      ProcessValue <- "F_Descargador_No"
   GraphicIOField "Campo ES gráfico_18" at 1195,401 size 28x28; PictureList "CheckBox"
      ProcessValue <- "F_Referencia_Menor_Descargador"
   IOField "Campo ES_7" at 1018,73 size 80x32; FormatPattern 9999999; Unit  mm
      ProcessValue <- "PosiciónEspera_F(Ant)"
   IOField "Campo ES_8" at 1018,97 size 80x32; FormatPattern 9999999; Unit  mm
      ProcessValue <- "PosiciónE1H1_F(Ant)"
   IOField "Campo ES_9" at 1018,121 size 80x32; FormatPattern 9999999; Unit  mm
      ProcessValue <- "PosiciónE1H2_F(Ant)"
   IOField "Campo ES_10" at 1018,145 size 80x32; FormatPattern 9999999; Unit  mm
      ProcessValue <- "PosiciónE2H1_F(Ant)"
   IOField "Campo ES_12" at 1018,169 size 80x32; FormatPattern 9999999; Unit  mm
      ProcessValue <- "PosiciónE2H2_F(Ant)"
   IOField "Campo ES_13" at 1018,193 size 80x32; FormatPattern 9999999; Unit  mm
      ProcessValue <- "PosiciónEntrega_F(Ant)"
   TextField "Campo de texto_34" at 249,678 size 130x18; Text 'DATOS PIEZA ACTUAL'
   TextField "Campo de texto_35" at 403,678 size 12x18; Text 'A'
   IOField "Champ E/S_24" at 414,675 size 53x25; FormatPattern 9999999
      ProcessValue <- "Pinza\Pinza.A"
      Appearance <- "Pinza\Pinza.PresenciaPieza"
   IOField "Champ E/S_25" at 483,675 size 53x25; FormatPattern 9999999
      ProcessValue <- "Pinza\Pinza.B"
      Appearance <- "Pinza\Pinza.PresenciaPieza"
   IOField "Champ E/S_26" at 554,675 size 53x24; FormatPattern 9999999
      ProcessValue <- "Pinza\Pinza.C"
      Appearance <- "Pinza\Pinza.PresenciaPieza"
   IOField "Champ E/S_27" at 629,675 size 53x25; FormatPattern 9999999
      ProcessValue <- "Pinza\Pinza.D"
      Appearance <- "Pinza\Pinza.PresenciaPieza"
   TextField "Campo de texto_36" at 472,678 size 11x18; Text 'B'
   TextField "Campo de texto_37" at 541,678 size 11x18; Text 'C'
   TextField "Campo de texto_38" at 616,678 size 12x18; Text 'D'
   TextField "Campo de texto_32" at 696,37 size 42x23; Text 'Pinza'
   TextField "Template_Plantilla_Campo de texto_4" at 696,67 size 568x3; Text 'Text'
   TextField "Template_Plantilla_Campo de texto_1" at 696,439 size 568x3; Text 'Text'
   TextField "Campo de texto_7" at 947,396 size 82x36; Text 'MOVIMIENTO SEGURO'
      Visibility <- "F_MovimientoSeguro"
      Appearance <- "F_MovimientoSeguro"
   TextField "Campo de texto_33" at 726,368 size 87x33; Text 'Tenaza Pleg. Atrás'
   TextField "Campo de texto_39" at 815,368 size 63x33; Text 'Herr. 1 OFF'
   TextField "Template_Plantilla_Campo de texto_3" at 696,359 size 568x3; Text 'Text'
   TextField "Campo de texto_43" at 882,368 size 63x33; Text 'Herr. 2 OFF'
   TextField "Campo de texto_18" at 1072,368 size 95x33; Text 'Descargador Atrás'
   TextField "Campo de texto_19" at 1160,368 size 95x33; Text 'Movimiento Corto'
   TextField "Campo de texto_10" at 719,242 size 191x25; Text 'Escalador relación mecánica'
   TextField "Campo de texto_13" at 719,262 size 191x25; Text 'Offset mecánico'
   TextField "Campo de texto_20" at 949,556 size 41x18; Text 'Martillo'
      Visibility <- "MANU"
   TextField "Campo de texto_23" at 825,556 size 35x18; Text 'Matriz'
      Visibility <- "MANU"
   TextField "Campo de texto_42" at 737,581 size 42x18; Text 'Herr. 1'
      Visibility <- "MANU"
   TextField "Campo de texto_45" at 737,622 size 42x18; Text 'Herr. 2'
      Visibility <- "MANU"
   TextField "Campo de texto_44" at 739,471 size 31x18; Text 'Pinza'
      Visibility <- "MANU"
   GraphicView "Visor de gráficos_1" at 1047,570 size 74x43; Picture "EMR2"
      Visibility <- "MANU"
   GraphicView "Visor de gráficos_2" at 1048,612 size 74x43; Picture "F1-3 EMR2"
      Visibility <- "MANU"
   GraphicView "Visor de gráficos_3" at 1152,612 size 74x43; Picture "F2-4 EMR2"
      Visibility <- "MANU"
   GraphicView "Visor de gráficos_4" at 1150,570 size 74x43; Picture "F1-3 EMR2"
      Visibility <- "MANU"
   GraphicView "Visor de gráficos_5" at 1126,590 size 12x12; Picture "outline_arrow_forward_ios_white_18dp"
      Visibility <- "MANU"
   GraphicView "Visor de gráficos_6" at 1135,590 size 12x12; Picture "outline_arrow_forward_ios_white_18dp"
      Visibility <- "MANU"
   GraphicView "Visor de gráficos_7" at 1126,632 size 12x12; Picture "outline_arrow_forward_ios_white_18dp"
      Visibility <- "MANU"
   GraphicView "Visor de gráficos_8" at 1135,632 size 12x12; Picture "outline_arrow_forward_ios_white_18dp"
      Visibility <- "MANU"
   TextField "Campo de texto_40" at 740,522 size 134x18; Text 'Bloque de Herramientas'
      Visibility <- "MANU"
   Button "Botón_42" at 48,625 size 40x40; TextOff 'Vista Condiciones'; PictureOff "Gráfico_7"
      on Click: ActivateScreen("eProC - 10 - Estados F_HW", 0)
   Button "Botón_11" at 1224,27 size 40x37; TextOff 'Vista Condiciones'; PictureOff "Tool"; Authorization "Nivel 3"
      on Click: ActivateScreen("eProC - 11 Referencias F-PL", 0)
   Button "Template_Plantilla_Bouton_2" at 1085,715 size 193x53; TextOff 'ALARMAS / DEFAUT'
      on Press: ActivateScreen("eProC - Alarmas", 0)
      Visibility <- "DB_OP.P_DEFAUT"

screen "eProC - 10 - Estados F_HW" 1280x768, template "Template"
   GraphicIOField "Campo ES gráfico_6" at 554,292 size 718x282; PictureList "Grupo 3 - Pinza1"
      ProcessValue <- "Alarma_Pinza"
   Polygon "Polígono_2" at 281,432 size 517x163
      Visibility <- "Pinza\Pinza.PresenciaPieza"
   Circle "Cercle_16" at 798,434 size 10x10
      Appearance <- "29S4"
   TextField "Campo de texto_29" at 910,349 size 114x18; Text '29S4 - Pinza Abierta'
   TextField "Campo de texto_30" at 894,313 size 116x18; Text '29S5 - Pinza Cerrada'
   Circle "Cercle_17" at 798,418 size 10x10
      Appearance <- "29S5"
   GraphicIOField "Campo ES gráfico_8" at 192,179 size 289x268; PictureList "Formador"
      ProcessValue <- "Alarma_Formador"
   Circle "Cercle_6" at 331,217 size 10x10
      Appearance <- "28S5"
   Circle "Cercle_7" at 331,246 size 10x10
      Appearance <- "28S6"
   TextField "Campo de texto_3" at 54,201 size 180x18; Text '28S5 - Herramientas Bloqueadas'
   TextField "Campo de texto_5" at 36,229 size 200x18; Text '28S6 - Herramientas Desbloqueadas'
   Circle "Cercle_8" at 406,291 size 10x10
      Appearance <- "28S3"
   Circle "Cercle_9" at 418,306 size 10x10
      Appearance <- "28S4"
   Circle "Cercle_10" at 460,360 size 10x10
      Appearance <- "28S1"
   Circle "Cercle_1" at 437,332 size 10x10
      Appearance <- "28S2"
   Circle "Cercle_0" at 371,397 size 10x10
      Appearance <- "27S5"
   Circle "Cercle_2" at 348,367 size 10x10
      Appearance <- "27S6"
   Circle "Cercle_18" at 313,326 size 10x10
      Appearance <- "27S7"
   Circle "Cercle_19" at 326,344 size 10x10
      Appearance <- "27S8"
   TextField "Campo de texto_10" at 488,240 size 146x18; Text '28S3 - Herr. 2 Matriz OFF'
   TextField "Campo de texto_15" at 496,267 size 142x18; Text '28S4 - Herr. 2 Matriz ON'
   TextField "Campo de texto_16" at 522,323 size 152x18; Text '28S1 - Herr. 2 Martillo OFF'
   TextField "Campo de texto_17" at 506,295 size 148x18; Text '28S2 - Herr. 2 Martillo ON'
   TextField "Campo de texto_11" at 44,381 size 146x18; Text '27S7 - Herr. 1 Matriz OFF'
   TextField "Campo de texto_19" at 46,411 size 142x18; Text '27S8 - Herr. 1 Matriz ON'
   TextField "Campo de texto_20" at 73,488 size 152x18; Text '27S5 - Herr. 1 Martillo OFF'
   TextField "Campo de texto_21" at 58,452 size 148x18; Text '27S6 - Herr. 1 Martillo ON'
   Button "Botón_42" at 48,625 size 40x40; TextOff 'Vista Condiciones'; PictureOff "Gráfico_6"
      on Click: ActivateScreen("eProC - 10 - Estados F", 0)
   TextField "Campo de texto_1" at 804,90 size 41x18; Text 'Martillo'
      Visibility <- "MANU"
   TextField "Campo de texto_23" at 680,90 size 35x18; Text 'Matriz'
      Visibility <- "MANU"
   TextField "Campo de texto_42" at 592,115 size 42x18; Text 'Herr. 1'
      Visibility <- "MANU"
   TextField "Campo de texto_45" at 592,156 size 42x18; Text 'Herr. 2'
      Visibility <- "MANU"
   TextField "Campo de texto_44" at 732,638 size 31x18; Text 'Pinza'
      Visibility <- "MANU"
   GraphicView "Visor de gráficos_1" at 904,108 size 74x43; Picture "EMR2"
      Visibility <- "MANU"
   GraphicView "Visor de gráficos_2" at 905,150 size 74x43; Picture "F1-3 EMR2"
      Visibility <- "MANU"
   GraphicView "Visor de gráficos_3" at 1009,150 size 74x43; Picture "F2-4 EMR2"
      Visibility <- "MANU"
   GraphicView "Visor de gráficos_4" at 1007,108 size 74x43; Picture "F1-3 EMR2"
      Visibility <- "MANU"
   GraphicView "Visor de gráficos_5" at 983,128 size 12x12; Picture "outline_arrow_forward_ios_white_18dp"
      Visibility <- "MANU"
   GraphicView "Visor de gráficos_6" at 992,128 size 12x12; Picture "outline_arrow_forward_ios_white_18dp"
      Visibility <- "MANU"
   GraphicView "Visor de gráficos_7" at 983,170 size 12x12; Picture "outline_arrow_forward_ios_white_18dp"
      Visibility <- "MANU"
   GraphicView "Visor de gráficos_8" at 992,170 size 12x12; Picture "outline_arrow_forward_ios_white_18dp"
      Visibility <- "MANU"
   TextField "Campo de texto_40" at 270,118 size 134x18; Text 'Bloque de Herramientas'
      Visibility <- "MANU"
   Button "Template_Plantilla_Bouton_2" at 1085,715 size 193x53; TextOff 'ALARMAS / DEFAUT'
      on Press: ActivateScreen("eProC - Alarmas", 0)
      Visibility <- "DB_OP.P_DEFAUT"
   TextField "Campo de texto_12" at 460,410 size 81x18; Text 'Herramienta 2'
   TextField "Campo de texto_13" at 366,434 size 81x18; Text 'Herramienta 1'
   Button "Botón_6" at 772,630 size 58x33; TextOff 'Avance'
      on Press: SetTag("DB_OP.RC2", 31); SetBit("DB_OP.OP_SELMANU2")
      Visibility <- "MANU"
      Appearance <- "DB_OP.RC2"
   Button "Botón_7" at 827,630 size 58x33; TextOff 'Retroc.'
      on Press: SetTag("DB_OP.RC2", 32); SetBit("DB_OP.OP_SELMANU2")
      Visibility <- "MANU"
      Appearance <- "DB_OP.RC2"
   Button "Botón_8" at 903,630 size 58x33; TextOff 'Abrir'
      on Press: SetTag("DB_OP.RC2", 33); SetBit("DB_OP.OP_SELMANU2")
      Visibility <- "MANU"
      Appearance <- "DB_OP.RC2"
   Button "Botón_9" at 959,630 size 58x33; TextOff 'Cerrar'
      on Press: SetTag("DB_OP.RC2", 34); SetBit("DB_OP.OP_SELMANU2")
      Visibility <- "MANU"
      Appearance <- "DB_OP.RC2"
   Button "Botón_34" at 496,110 size 58x33; TextOff 'Bajar'
      on Press: SetTag("DB_OP.RC2", 40); SetBit("DB_OP.OP_SELMANU2")
      Visibility <- "MANU"
      Appearance <- "DB_OP.RC2"
   Button "Botón_35" at 439,110 size 58x33; TextOff 'Subir'
      on Press: SetTag("DB_OP.RC2", 41); SetBit("DB_OP.OP_SELMANU2")
      Visibility <- "MANU"
      Appearance <- "DB_OP.RC2"
   Button "Botón_20" at 765,110 size 58x33; TextOff 'ON'
      on Press: SetTag("DB_OP.RC2", 42); SetBit("DB_OP.OP_SELMANU2")
      Visibility <- "MANU"
      Appearance <- "DB_OP.RC2"
   Button "Botón_21" at 765,149 size 58x33; TextOff 'ON'
      on Press: SetTag("DB_OP.RC2", 46); SetBit("DB_OP.OP_SELMANU2")
      Visibility <- "MANU"
      Appearance <- "DB_OP.RC2"
   Button "Botón_22" at 821,110 size 58x33; TextOff 'OFF'
      on Press: SetTag("DB_OP.RC2", 43); SetBit("DB_OP.OP_SELMANU2")
      Visibility <- "MANU"
      Appearance <- "DB_OP.RC2"
   Button "Botón_23" at 821,149 size 58x33; TextOff 'OFF'
      on Press: SetTag("DB_OP.RC2", 47); SetBit("DB_OP.OP_SELMANU2")
      Visibility <- "MANU"
      Appearance <- "DB_OP.RC2"
   Button "Botón_28" at 641,110 size 58x33; TextOff 'ON'
      on Press: SetTag("DB_OP.RC2", 44); SetBit("DB_OP.OP_SELMANU2")
      Visibility <- "MANU"
      Appearance <- "DB_OP.RC2"
   Button "Botón_5" at 641,148 size 58x33; TextOff 'ON'
      on Press: SetTag("DB_OP.RC2", 48); SetBit("DB_OP.OP_SELMANU2")
      Visibility <- "MANU"
      Appearance <- "DB_OP.RC2"
   Button "Botón_10" at 697,110 size 58x33; TextOff 'OFF'
      on Press: SetTag("DB_OP.RC2", 45); SetBit("DB_OP.OP_SELMANU2")
      Visibility <- "MANU"
      Appearance <- "DB_OP.RC2"
   Button "Botón_31" at 697,148 size 58x33; TextOff 'OFF'
      on Press: SetTag("DB_OP.RC2", 49); SetBit("DB_OP.OP_SELMANU2")
      Visibility <- "MANU"
      Appearance <- "DB_OP.RC2"

screen "eProC - 11 Referencias F-PL" 1280x768, template "Template"
   GraphicView "Visor de gráficos_1" at 134,72 size 979x505; Picture "Referencias"
   IOField "Champ E/S" at 340,310 size 80x27; Authorization "Nivel 2"; FormatPattern 9999999
      ProcessValue <- "Distancia_entre_Herramienta1_y_Pos0_F"
   IOField "Champ E/S_0" at 540,342 size 80x26; Authorization "Nivel 2"; FormatPattern 9999999
      ProcessValue <- "Distancia_entre_Pos0_y_Tenaza_F"
   TextField "Campo de texto_1" at 334,240 size 90x68; Text 'Distancia de Herramienta 1 a posición 0mm Pinza'
   TextField "Campo de texto_3" at 526,300 size 126x36; Text 'Distancia 0mm Pinza a Tenaza Plegadora'
   IOField "Champ E/S_2" at 552,526 size 80x26; Authorization "Nivel 2"; FormatPattern 9999999
      ProcessValue <- "Distancia_entre_Pos0_y_Descargador_F"
   TextField "Campo de texto_6" at 505,553 size 176x36; Text 'Distancia posición 0mm Pinza al Descargador'
   IOField "Champ E/S_3" at 235,566 size 80x27; Authorization "Nivel 2"; FormatPattern 9999999
      ProcessValue <- "Distancia_entre_Herramientas_F"
   TextField "Campo de texto_7" at 230,594 size 93x36; Text 'Distancia entre Herramientas'
   IOField "Champ E/S_4" at 592,610 size 80x26; Authorization "Nivel 2"; FormatPattern s9999999999
      ProcessValue <- "PosiciónMáxima_F"
   TextField "Campo de texto_8" at 587,636 size 93x36; Text 'Distancia Avance Máximo'
   IOField "Champ E/S_1" at 907,300 size 80x26; Authorization "Nivel 2"; FormatPattern 9999999
      ProcessValue <- "Distancia_entre_Pleg_Alin_PL"
   TextField "Campo de texto_2" at 861,330 size 196x20; Text 'Distancia de Plegador a Alineador'
   Switch "Interruptor_1" at 209,115 size 125x80; TextOn 'SI'; CaptionText 'Habilitar reglas'; TextOff 'NO'
      ProcessValue <- "HabilitarReglasBaluff"
   Button "Botón_1" at 440,76 size 135x50; TextOff 'Referenciar PL1'
      on Release: ResetBit("SolRef_PL1")
      on Press: SetBit("SolRef_PL1")
      Appearance <- "Homing_PL1"
      ObjectEnable <- "HabRefPleg"
      Visibility <- "HabRefPleg"
   Button "Botón_2" at 941,76 size 135x50; TextOff 'Referenciar PL2'
      on Release: ResetBit("SolRef_PL2")
      on Press: SetBit("SolRef_PL2")
      Appearance <- "Homing_PL2"
      ObjectEnable <- "HabRefPleg"
      Visibility <- "HabRefPleg"
   Button "Template_Plantilla_Bouton_2" at 1085,715 size 193x53; TextOff 'ALARMAS / DEFAUT'
      on Press: ActivateScreen("eProC - Alarmas", 0)
      Visibility <- "DB_OP.P_DEFAUT"

screen "eProC - Recetas" 1280x768, template "Template"
   IOField "Champ E/S_43" at 357,162 size 98x23; FormatPattern 9999999; Unit  mm
      ProcessValue <- "Receta\Recetas.B"
   IOField "Champ E/S_44" at 869,304 size 90x23; FormatPattern 9999999; Unit  mm
      ProcessValue <- "Receta\Recetas.C"
   IOField "Champ E/S_46" at 743,113 size 96x24; FormatPattern s999999; Unit  mm
      ProcessValue <- "Receta\Recetas.F2"
   IOField "Champ E/S_47" at 743,90 size 90x23; FormatPattern s999999; Unit  mm
      ProcessValue <- "Receta\Recetas.F1"
   IOField "Champ E/S_48" at 561,90 size 94x23; FormatPattern s999999; Unit  mm
      ProcessValue <- "Receta\Recetas.F3"
   IOField "Champ E/S_49" at 581,137 size 96x24; FormatPattern s999999; Unit  mm
      ProcessValue <- "Receta\Recetas.PL1_2"
   IOField "Champ E/S_50" at 193,137 size 91x24; FormatPattern s999999; Unit  mm
      ProcessValue <- "Receta\Recetas.PL1_1"
   IOField "Champ E/S_51" at 1165,137 size 94x24; FormatPattern s999999; Unit  mm
      ProcessValue <- "Receta\Recetas.PL2_1"
   TextField "Campo de texto_56" at 340,160 size 17x26; Text 'B'
   TextField "Campo de texto_57" at 852,302 size 17x26; Text 'C'
   IOField "Champ E/S_52" at 1121,303 size 88x24; FormatPattern 9999999; Unit  mm
      ProcessValue <- "Receta\Recetas.D"
   TextField "Campo de texto_60" at 1103,302 size 19x26; Text 'D'
   IOField "Champ E/S_53" at 561,112 size 94x25; FormatPattern s999999; Unit  mm
      ProcessValue <- "Receta\Recetas.F4"
   IOField "Champ E/S_54" at 764,137 size 93x24; FormatPattern s999999; Unit  mm
      ProcessValue <- "Receta\Recetas.PL2_2"
   TextField "Campo de texto_62" at 556,302 size 17x26; Text 'A'
   IOField "Champ E/S_55" at 575,304 size 94x23; FormatPattern 9999999; Unit  mm
      ProcessValue <- "Receta\Recetas.A"
   TextField "Campo de texto_63" at 542,138 size 40x22; Text 'PL1-2'
   TextField "Campo de texto_64" at 726,113 size 20x22; Text 'F2'
   TextField "Campo de texto_65" at 152,138 size 40x22; Text 'PL1-1'
   TextField "Campo de texto_66" at 726,89 size 20x22; Text 'F1'
   TextField "Campo de texto_67" at 725,138 size 40x22; Text 'PL2-2'
   TextField "Campo de texto_68" at 541,113 size 20x22; Text 'F4'
   TextField "Campo de texto_69" at 1124,138 size 40x22; Text 'PL2-1'
   TextField "Campo de texto_70" at 541,89 size 20x22; Text 'F3'
   RecipeView "RecipeView" at 25,65 size 307x64; RecipeNameCaption 'Receta:'; DataRecordNameCaption 'Receta:'; ValueCaption 'Valor'; RecipeNrCaption 'N.º:'; DataRecordNrCaption 'Nº:'; EntryNameCaption 'Nombre de entrada'; Recipe "Pieza"; Tag4DataRecord "Receta\Recetas.Nombre"
   Button "Button_7" at 856,371 size 82x33; TextOff 'Cargar'; PictureOff "Flèche_Droite"
      on Press: SetBit("Receta\Recetas.x_M2"); function_eba64363('REFERENCE', "Receta\Recetas.Nombre", 1, N)
      Appearance <- "Receta\Recetas.x_M2"
   TextField "Campo de texto_15" at 953,376 size 72x22; Text 'Almacén 2'
   IOField "Champ E/S_57" at 1041,376 size 118x24; FormatPattern ????????????????????
      ProcessValue <- "Almacén 2\PAlmacén.Nombre"
   TextField "Campo de texto_59" at 39,37 size 159x26; Text 'Selección de Receta'
   Button "Button_6" at 42,368 size 82x35; TextOff 'Cargar'; PictureOff "Flèche_Droite"
      on Press: SetBit("Receta\Recetas.x_M1"); function_eba64363('REFERENCE', "Receta\Recetas.Nombre", 1, N)
      Appearance <- "Receta\Recetas.x_M1"
   TextField "Campo de texto_14" at 139,375 size 72x22; Text 'Almacén 1'
   IOField "Champ E/S_56" at 227,375 size 120x24; FormatPattern ????????????????????
      ProcessValue <- "Almacén 1\PAlmacén.Nombre"
   IOField "Champ E/S_1" at 289,304 size 90x23; FormatPattern 9999999; Unit  mm
      ProcessValue <- "Receta\Recetas.C"
   TextField "Campo de texto_1" at 272,302 size 17x26; Text 'C'
   IOField "Champ E/S_2" at 41,303 size 88x24; FormatPattern 9999999; Unit  mm
      ProcessValue <- "Receta\Recetas.D"
   TextField "Campo de texto_2" at 23,302 size 19x26; Text 'D'
   Button "Template_Plantilla_Bouton_1" at 345,50 size 150x63; TextOff 'EDITAR RECETAS / SYSTEM'; Authorization "Nivel 3"
      on Click: ActivateScreen("eProC - Edición Recetas", 0)
   Button "Template_Plantilla_Botón_32" at 129,715 size 150x53; TextOff 'SELECCIÓN RECETAS'
   Button "Template_Plantilla_Bouton_2" at 1085,715 size 193x53; TextOff 'ALARMAS / DEFAUT'
      on Press: ActivateScreen("eProC - Alarmas", 0)
      Visibility <- "DB_OP.P_DEFAUT"
   IOField "Campo ES_1" at 321,415 size 130x34; FormatPattern 9999999999
      ProcessValue <- "Descargador-ID_Bobina_Alm1"
   IOField "Campo ES_2" at 1136,415 size 130x34; FormatPattern 9999999999
      ProcessValue <- "Descargador-ID_Bobina_Alm2"
   DateTimeField "Campo de fecha y hora_1" at 180,415 size 131x34
      ProcessValue <- "Descargador-FechaCorte_Alm1"
   DateTimeField "Campo de fecha y hora_2" at 995,415 size 131x34
      ProcessValue <- "Descargador-FechaCorte_Alm2"
   SymbolicIOField "Campo ES simbólico_1" at 41,415 size 130x34; TextOff '0'; TextOn '1'; TextList "Proveedor"
      ProcessValue <- "Proveedor_Indexado_Alm1"
   SymbolicIOField "Campo ES simbólico_2" at 856,415 size 130x34; TextOff '0'; TextOn '1'; TextList "Proveedor"
      ProcessValue <- "Proveedor_Indexado_Alm2"
   IOField "Champ E/S_74" at 302,520 size 64x32; Authorization "Nivel 1"; FormatPattern s999999; Unit   
      ProcessValue <- "Almacén 1\PAlmacén.F2"
   IOField "Champ E/S_75" at 302,493 size 64x32; Authorization "Nivel 1"; FormatPattern s999999; Unit   
      ProcessValue <- "Almacén 1\PAlmacén.F1"
   IOField "Champ E/S_76" at 86,498 size 64x32; Authorization "Nivel 1"; FormatPattern s999999; Unit   
      ProcessValue <- "Almacén 1\PAlmacén.F3"
   IOField "Champ E/S_77" at 86,471 size 64x32; Authorization "Nivel 1"; FormatPattern s999999; Unit   
      ProcessValue <- "Almacén 1\PAlmacén.PL1_2"
   IOField "Champ E/S_78" at 86,648 size 64x32; Authorization "Nivel 1"; FormatPattern s999999; Unit   
      ProcessValue <- "Almacén 1\PAlmacén.PL1_1"
   IOField "Champ E/S_79" at 302,651 size 64x32; Authorization "Nivel 1"; FormatPattern s999999; Unit   
      ProcessValue <- "Almacén 1\PAlmacén.PL2_1"
   IOField "Champ E/S_81" at 86,525 size 64x32; Authorization "Nivel 1"; FormatPattern s999999; Unit   
      ProcessValue <- "Almacén 1\PAlmacén.F4"
   IOField "Champ E/S_82" at 302,466 size 64x32; Authorization "Nivel 1"; FormatPattern s999999; Unit   
      ProcessValue <- "Almacén 1\PAlmacén.PL2_2"
   TextField "Campo de texto_80" at 46,476 size 40x22; Text 'PL1-2'
   TextField "Campo de texto_81" at 366,526 size 20x22; Text 'F2'
   TextField "Campo de texto_82" at 46,652 size 40x22; Text 'PL1-1'
   TextField "Campo de texto_83" at 366,497 size 20x22; Text 'F1'
   TextField "Campo de texto_84" at 364,471 size 40x22; Text 'PL2-2'
   TextField "Campo de texto_85" at 66,531 size 20x22; Text 'F4'
   TextField "Campo de texto_86" at 364,655 size 40x22; Text 'PL2-1'
   TextField "Campo de texto_87" at 66,502 size 20x22; Text 'F3'
   IOField "Champ E/S_15" at 904,498 size 64x32; Authorization "Nivel 1"; FormatPattern s999999; Unit   
      ProcessValue <- "Almacén 2\PAlmacén.F3"
   IOField "Champ E/S_16" at 904,471 size 64x32; Authorization "Nivel 1"; FormatPattern s999999; Unit   
      ProcessValue <- "Almacén 2\PAlmacén.PL1_2"
   IOField "Champ E/S_58" at 904,648 size 65x32; Authorization "Nivel 1"; FormatPattern s999999; Unit   
      ProcessValue <- "Almacén 2\PAlmacén.PL1_1"
   IOField "Champ E/S_60" at 904,525 size 64x32; Authorization "Nivel 1"; FormatPattern s999999; Unit   
      ProcessValue <- "Almacén 2\PAlmacén.F4"
   TextField "Campo de texto_53" at 865,476 size 40x22; Text 'PL1-2'
   TextField "Campo de texto_55" at 865,652 size 40x22; Text 'PL1-1'
   TextField "Campo de texto_58" at 885,531 size 20x22; Text 'F4'
   TextField "Campo de texto_7" at 885,502 size 20x22; Text 'F3'
   IOField "Champ E/S_13" at 1119,520 size 64x32; Authorization "Nivel 1"; FormatPattern s999999; Unit   
      ProcessValue <- "Almacén 2\PAlmacén.F2"
   IOField "Champ E/S_14" at 1119,493 size 64x32; Authorization "Nivel 1"; FormatPattern s999999; Unit   
      ProcessValue <- "Almacén 2\PAlmacén.F1"
   IOField "Champ E/S_59" at 1119,651 size 64x32; Authorization "Nivel 1"; FormatPattern s999999; Unit   
      ProcessValue <- "Almacén 2\PAlmacén.PL2_1"
   IOField "Champ E/S_61" at 1119,466 size 64x32; Authorization "Nivel 1"; FormatPattern s999999; Unit   
      ProcessValue <- "Almacén 2\PAlmacén.PL2_2"
   TextField "Campo de texto_54" at 1180,526 size 20x22; Text 'F2'
   TextField "Campo de texto_4" at 1180,497 size 20x22; Text 'F1'
   TextField "Campo de texto_5" at 1180,471 size 40x22; Text 'PL2-2'
   TextField "Campo de texto_6" at 1180,655 size 40x22; Text 'PL2-1'
   IOField "Champ E/S_3" at 86,581 size 64x32; Authorization "Nivel 1"; FormatPattern s999999; Unit   
      ProcessValue <- "Almacén 1\PAlmacén.C"
   TextField "Campo de texto_3" at 66,587 size 13x22; Text 'C'
   IOField "Champ E/S_4" at 904,581 size 64x32; Authorization "Nivel 1"; FormatPattern s999999; Unit   
      ProcessValue <- "Almacén 2\PAlmacén.C"
   TextField "Campo de texto_8" at 885,587 size 13x22; Text 'C'

screen "eProC - Defectos" 1280x768, template "Template"
   TextField "Campo de texto_14" at 18,389 size 97x28; Text 'Almacén 2'
   TextField "Campo de texto_7" at 693,45 size 95x28; Text 'Esquina 1'
   TextField "Campo de texto_8" at 532,45 size 95x28; Text 'Esquina 2'
   TextField "Campo de texto_9" at 364,97 size 138x28; Text 'Herramienta 1'
   TextField "Campo de texto_10" at 364,154 size 138x28; Text 'Herramienta 2'
   TextField "Campo de texto_2" at 982,66 size 85x28; Text 'Contador'
   TextField "Campo de texto_1" at 18,45 size 97x28; Text 'Almacén 1'
   TextField "Campo de texto_3" at 693,381 size 90x28; Text 'Esquina 1'
   TextField "Campo de texto_4" at 532,381 size 90x28; Text 'Esquina 2'
   TextField "Campo de texto_5" at 364,433 size 133x28; Text 'Herramienta 1'
   TextField "Campo de texto_6" at 364,490 size 133x28; Text 'Herramienta 2'
   TextField "Campo de texto_16" at 982,402 size 85x28; Text 'Contador'
   TextField "Campo de texto_11" at 316,306 size 102x28; Text 'Plegadores'
   TextField "Campo de texto_12" at 316,642 size 102x28; Text 'Plegadores'
   Button "Template_Plantilla_Botón_55" at 789,715 size 150x53; TextOff 'ACUSAR DEFECTO'
   IOField "Campo ES_1" at 980,106 size 96x32; FormatPattern 9999
      ProcessValue <- "Contador_def_Alm1"
   Button "Botón_1" at 520,92 size 120x40; TextOff 'E2 H1'
      on Click: function_dd21b452("Contador_def_Alm1", 1); SetTag("Defecto_Alm1", 3)
   Button "Botón_2" at 680,92 size 120x40; TextOff 'E1 H1'
      on Click: function_dd21b452("Contador_def_Alm1", 1); SetTag("Defecto_Alm1", 1)
   Button "Botón_3" at 520,148 size 120x40; TextOff 'E2 H2'
      on Click: function_dd21b452("Contador_def_Alm1", 1); SetTag("Defecto_Alm1", 4)
   Button "Botón_4" at 680,148 size 120x40; TextOff 'E1 H2'
      on Click: function_dd21b452("Contador_def_Alm1", 1); SetTag("Defecto_Alm1", 2)
   Button "Botón_5" at 472,300 size 120x40; TextOff 'PL1-2'
      on Click: function_dd21b452("Contador_def_Alm1", 1); SetTag("Defecto_Alm1", 5)
   Button "Botón_6" at 632,300 size 120x40; TextOff 'PL2-2'
      on Click: function_dd21b452("Contador_def_Alm1", 1); SetTag("Defecto_Alm1", 6)
   Button "Botón_7" at 980,146 size 120x40; TextOff 'Reset'
      on Click: SetTag("Contador_def_Alm1", 0)
   IOField "Campo ES_2" at 980,442 size 96x32; FormatPattern 9999
      ProcessValue <- "Contador_def_Alm2"
   Button "Botón_8" at 520,428 size 120x40; TextOff 'E2 H1'
      on Click: function_dd21b452("Contador_def_Alm2", 1); SetTag("Defecto_Alm2", 3)
   Button "Botón_9" at 680,428 size 120x40; TextOff 'E1 H1'
      on Click: function_dd21b452("Contador_def_Alm2", 1); SetTag("Defecto_Alm2", 1)
   Button "Botón_10" at 520,484 size 120x40; TextOff 'E2 H2'
      on Click: function_dd21b452("Contador_def_Alm2", 1); SetTag("Defecto_Alm2", 4)
   Button "Botón_11" at 680,484 size 120x40; TextOff 'E1 H2'
      on Click: function_dd21b452("Contador_def_Alm2", 1); SetTag("Defecto_Alm2", 2)
   Button "Botón_12" at 472,636 size 120x40; TextOff 'PL1-2'
      on Click: function_dd21b452("Contador_def_Alm2", 1); SetTag("Defecto_Alm2", 5)
   Button "Botón_13" at 632,636 size 120x40; TextOff 'PL2-2'
      on Click: function_dd21b452("Contador_def_Alm2", 1); SetTag("Defecto_Alm2", 6)
   Button "Botón_14" at 980,482 size 120x40; TextOff 'Reset'
      on Click: SetTag("Contador_def_Alm2", 0)
   Button "Template_Plantilla_Bouton_2" at 1085,715 size 193x53; TextOff 'ALARMAS / DEFAUT'
      on Press: ActivateScreen("eProC - Alarmas", 0)
      Visibility <- "DB_OP.P_DEFAUT"
   IOField "Champ E/S_1" at 122,392 size 171x24; FormatPattern ????????????????????
      ProcessValue <- "Almacén 2\PAlmacén.Nombre"
   IOField "Champ E/S_2" at 122,48 size 170x24; FormatPattern ????????????????????
      ProcessValue <- "Almacén 1\PAlmacén.Nombre"

VB script "Script_1"
   'NOTE : Appuyez sur <Ctrl><Espacement> pour lancer le script et afficher le large éventail de fonctions.
   'Ecrivez vos scripts en utilisant les fonctions système ou le modèle d'objet. Vous pouvez facilement accéder au
   'système via l'objet runtime IHM. Pour sélectionner rapidement une référence objet
   'vous pouvez appuyer sur <Alt><Flèche droite>. Vous pouvez créer des scripts complexes en ayant recours au
   'langage de programmation VBScript et accéder directement aux variables via le nom, par ex. tag = 5.
*)

(* ===== HMI "HMI_RT_2" =====
system functions are stored by id; their names below are inferred from use
connection "HMI_ServidorHTTP": Web, WebPanel

HMI tags "Tabla de variables estándar"
   "Descargador-PiezaPresente" : Bool AT Descargador-PiezaPresente, 1 s   // Unidad presente en el descargador (DB12DBX46.0)
   "31S1 (E8.0)" : Bool AT 31S1, 1 s   // Presencia Producto en Descargador
      on ChangeValue: "FuncionVB_1"()
   "Evento_ArchivarVariable_1" : Bool, internal   // Para guardar los datos del producto en almacen 1
      on ChangeValue: function_abcfba0d("Cota C_Alm1"); function_abcfba0d("Factor F1_Alm1"); function_abcfba0d("Factor F2_Alm1"); function_abcfba0d("Factor F3_Alm1"); function_abcfba0d("Factor F4_Alm1"); function_abcfba0d("Factor PL1-1_Alm1"); function_abcfba0d("Factor PL1-2_Alm1"); function_abcfba0d("Factor PL2-1_Alm1"); function_abcfba0d("Factor PL2-2_Alm1"); function_abcfba0d("ID_Proveedor_Alm1"); function_abcfba0d("ID_FechaCorte_Alm1"); function_abcfba0d("ID_Bobina_Alm1")
   "Evento_ArchivarVariable_2" : Bool, internal   // Para guardar lel posicionamiento de la pinza en almacen 1
      on ChangeValue: function_abcfba0d("PosReal_E1H1_Alm1"); function_abcfba0d("PosReal_E1H2_Alm1"); function_abcfba0d("PosReal_E2H1_Alm1"); function_abcfba0d("PosReal_E2H2_Alm1"); function_abcfba0d("PosReal_Entrega_Alm1"); function_abcfba0d("PosReal_Recepcion_Alm1"); function_abcfba0d("Consigna_E1H1_Alm1"); function_abcfba0d("Consigna_E1H2_Alm1"); function_abcfba0d("Consigna_E2H1_Alm1"); function_abcfba0d("Consigna_E2H2_Alm1"); function_abcfba0d("Consigna_Entrega_Alm1"); function_abcfba0d("Consigna_Recepcion_Alm1")
   "Evento_ArchivarVariable_3" : Bool, internal   // Para guardar el posicionamiento de los plegadores en almacen 1
      on ChangeValue: function_abcfba0d("PosiciónEntrega_PL1_A1"); function_abcfba0d("PosiciónEspera_PL1_A1"); function_abcfba0d("PosiciónPlegado1_PL1_A1"); function_abcfba0d("PosiciónPlegado2_PL1_A1"); function_abcfba0d("PosiciónRecepción_PL1_A1"); function_abcfba0d("PosiciónEntrega_PL2_A1"); function_abcfba0d("PosiciónEspera_PL2_A1"); function_abcfba0d("PosiciónPlegado1_PL2_A1"); function_abcfba0d("PosiciónPlegado2_PL2_A1"); function_abcfba0d("PosiciónRecepción_PL2_A1")
   "Descargador-Almacen" : Bool AT Descargador-Almacen, 1 s   // Si este bit es 0 la unidad proviene del almacén 1, si vale 1 del almacén 2 (DB12DBX46.1)
   "Evento_ArchivarVariable_4" : Bool, internal   // Para guardar los datos del producto en almacen 2
      on ChangeValue: function_abcfba0d("Cota C_Alm2"); function_abcfba0d("Factor F1_Alm2"); function_abcfba0d("Factor F2_Alm2"); function_abcfba0d("Factor F3_Alm2"); function_abcfba0d("Factor F4_Alm2"); function_abcfba0d("Factor PL1-1_Alm2"); function_abcfba0d("Factor PL1-2_Alm2"); function_abcfba0d("Factor PL2-1_Alm2"); function_abcfba0d("Factor PL2-2_Alm2"); function_abcfba0d("ID_Prov_Ind_Alm2"); function_abcfba0d("ID_FechaCorte_Alm2"); function_abcfba0d("ID_Bobina_Alm2")
   "Aux1" : Bool, internal   // utilizada en FuncionVB_1
   "Aux2" : Bool, internal   // para entrada de graficos en imagen ppal
   "Almacén 1\PAlmacén.Nombre" : String[10] AT Almacén 1\PAlmacén.Nombre, 1 min
   "Almacén 2\PAlmacén.Nombre" : String[10] AT Almacén 2\PAlmacén.Nombre, 1 min
   "Evento_ArchivarVariable_5" : Bool, internal   // Para guardar lel posicionamiento de la pinza en almacen 2
      on ChangeValue: function_abcfba0d("PosReal_E1H1_Alm2"); function_abcfba0d("PosReal_E1H2_Alm2"); function_abcfba0d("PosReal_E2H1_Alm2"); function_abcfba0d("PosReal_E2H2_Alm2"); function_abcfba0d("PosReal_Entrega_Alm2"); function_abcfba0d("PosReal_Recepcion_Alm2"); function_abcfba0d("Consigna_E1H1_Alm2"); function_abcfba0d("Consigna_E1H2_Alm2"); function_abcfba0d("Consigna_E2H1_Alm2"); function_abcfba0d("Consigna_E2H2_Alm2"); function_abcfba0d("Consigna_Entrega_Alm2"); function_abcfba0d("Consigna_Resepcion_Alm2")
   "Evento_ArchivarVariable_6" : Bool, internal   // Para guardar el posicionamiento de los plegadores en almacen 2
      on ChangeValue: function_abcfba0d("PosiciónEntrega_PL1_A2"); function_abcfba0d("PosiciónEntrega_PL2_A2"); function_abcfba0d("PosiciónEspera_PL1_A2"); function_abcfba0d("PosiciónEspera_PL2_A2"); function_abcfba0d("PosiciónPlegado1_PL1_A2"); function_abcfba0d("PosiciónPlegado1_PL2_A2"); function_abcfba0d("PosiciónPlegado2_PL1_A2"); function_abcfba0d("PosiciónPlegado2_PL2_A2"); function_abcfba0d("PosiciónRecepción_PL1_A2"); function_abcfba0d("PosiciónRecepción_PL2_A2")
   "Aux3" : Bool, internal   // para simular botones en imagen ppal
   "Defecto_Alm1" : Int AT Defecto_Alm1, 1 s
   "Defecto_Alm2" : Int AT Defecto_Alm2, 1 s
   "Contador_def_Alm1" : Int AT Contador_def_Alm1, 1 s
      on ChangeValue: function_abcfba0d("Defecto_Alm1")
   "Contador_def_Alm2" : Int AT Contador_def_Alm2, 1 s
      on ChangeValue: function_abcfba0d("Defecto_Alm2")
   "31S8 (E8.7)" : Bool AT 31S8, 1 s   // Presencia Producto en Descargador

HMI tags "DatProducto_A1"
   "Cota C_Alm1" : Int AT Descargador-C, 1 s
   "Factor F1_Alm1" : Int AT Descargador-F1, 1 s
   "Factor F2_Alm1" : Int AT Descargador-F2, 1 s
   "Factor F3_Alm1" : Int AT Descargador-F3, 1 s
   "Factor F4_Alm1" : Int AT Descargador-F4, 1 s
   "Factor PL1-1_Alm1" : Int AT Descargador-PL1_1, 1 s
   "Factor PL1-2_Alm1" : Int AT Descargador-PL1_2, 1 s
   "Factor PL2-1_Alm1" : Int AT Descargador-PL2_1, 1 s
   "Factor PL2-2_Alm1" : Int AT Descargador-PL2_2, 1 s
   "ID_Bobina_Alm1" : DInt AT Descargador-ID_Bobina_Alm1, 1 s
   "ID_Proveedor_Alm1" : Int AT Proveedor_Indexado_Alm1, 1 s
   "ID_FechaCorte_Alm1" : DateTime AT Descargador-FechaCorte_Alm1, 1 s

HMI tags "PosPinza_A1"
   "PosReal_E1H1_Alm1" : DInt AT Pos_E1H1(3), 1 s   // DB26
   "PosReal_E1H2_Alm1" : DInt AT Pos_E1H2(3), 1 s   // DB26
   "PosReal_E2H1_Alm1" : DInt AT Pos_E2H1(3), 1 s   // DB26
   "PosReal_E2H2_Alm1" : DInt AT Pos_E2H2(3), 1 s   // DB26
   "PosReal_Entrega_Alm1" : DInt AT Pos_Entrega(3), 1 s   // DB26
   "PosReal_Recepcion_Alm1" : DInt AT Pos_Recepcion(3), 1 s   // DB26
   "Consigna_E1H1_Alm1" : DInt AT PosiciónE1H1_F(Ant), 1 s   // DB18
   "Consigna_E1H2_Alm1" : DInt AT PosiciónE1H2_F(Ant), 1 s   // DB18
   "Consigna_E2H1_Alm1" : DInt AT PosiciónE2H1_F(Ant), 1 s   // DB18
   "Consigna_E2H2_Alm1" : DInt AT PosiciónE2H2_F(Ant), 1 s   // DB18
   "Consigna_Entrega_Alm1" : DInt AT PosiciónEntrega_F(Ant), 1 s   // DB18
   "Consigna_Recepcion_Alm1" : DInt AT PosiciónEspera_F(Ant), 1 s   // DB18

HMI tags "PosPlegadores_A1"
   "PosiciónEntrega_PL1_A1" : DInt AT PosiciónEntrega_PL1(Ant), 1 s   // DB57
   "PosiciónEntrega_PL2_A1" : DInt AT PosiciónEntrega_PL2(Ant), 1 s   // DB58
   "PosiciónEspera_PL1_A1" : DInt AT PosiciónEspera_PL1(Ant), 1 s   // DB57
   "PosiciónEspera_PL2_A1" : DInt AT PosiciónEspera_PL2(Ant), 1 s   // DB58
   "PosiciónPlegado1_PL1_A1" : DInt AT PosiciónPlegado1_PL1(Ant), 1 s   // DB57
   "PosiciónPlegado1_PL2_A1" : DInt AT PosiciónPlegado1_PL2(Ant), 1 s   // DB58
   "PosiciónPlegado2_PL1_A1" : DInt AT PosiciónPlegado2_PL1(Ant), 1 s   // DB57
   "PosiciónPlegado2_PL2_A1" : DInt AT PosiciónPlegado2_PL2(Ant), 1 s   // DB58
   "PosiciónRecepción_PL1_A1" : DInt AT PosiciónRecepción_PL1(Ant), 1 s   // DB57
   "PosiciónRecepción_PL2_A1" : DInt AT PosiciónRecepción_PL2(Ant), 1 s   // DB58

HMI tags "DatProducto_A2"
   "Cota C_Alm2" : Int AT Descargador-C, 1 s
   "Factor F1_Alm2" : Int AT Descargador-F1, 1 s
   "Factor F2_Alm2" : Int AT Descargador-F2, 1 s
   "Factor F3_Alm2" : Int AT Descargador-F3, 1 s
   "Factor F4_Alm2" : Int AT Descargador-F4, 1 s
   "Factor PL1-1_Alm2" : Int AT Descargador-PL1_1, 1 s
   "Factor PL1-2_Alm2" : Int AT Descargador-PL1_2, 1 s
   "Factor PL2-1_Alm2" : Int AT Descargador-PL1_2, 1 s
   "Factor PL2-2_Alm2" : Int AT Descargador-PL2_2, 1 s
   "ID_Prov_Ind_Alm2" : Int AT Proveedor_Indexado_Alm2, 1 s
   "ID_Bobina_Alm2" : DInt AT Descargador-ID_Bobina_Alm2, 1 s
   "ID_FechaCorte_Alm2" : DateTime AT Descargador-FechaCorte_Alm2, 1 s

HMI tags "PosPinza_A2"
   "PosReal_E1H1_Alm2" : DInt AT Pos_E1H1(3), 1 s   // DB26
   "PosReal_E1H2_Alm2" : DInt AT Pos_E1H2(3), 1 s   // DB26
   "PosReal_E2H1_Alm2" : DInt AT Pos_E2H1(3), 1 s   // DB26
   "PosReal_E2H2_Alm2" : DInt AT Pos_E2H2(3), 1 s   // DB26
   "PosReal_Entrega_Alm2" : DInt AT Pos_Entrega(3), 1 s   // DB26
   "PosReal_Recepcion_Alm2" : DInt AT Pos_Recepcion(3), 1 s   // DB26
   "Consigna_E1H1_Alm2" : DInt AT PosiciónE1H1_F(Ant), 1 s   // DB18
   "Consigna_E1H2_Alm2" : DInt AT PosiciónE1H2_F(Ant), 1 s   // DB18
   "Consigna_E2H1_Alm2" : DInt AT PosiciónE2H1_F(Ant), 1 s   // DB18
   "Consigna_E2H2_Alm2" : DInt AT PosiciónE2H2_F(Ant), 1 s   // DB18
   "Consigna_Entrega_Alm2" : DInt AT PosiciónEntrega_F(Ant), 1 s   // DB18
   "Consigna_Resepcion_Alm2" : DInt AT PosiciónEspera_F(Ant), 1 s   // DB18

HMI tags "PosPlegadores_A2"
   "PosiciónEntrega_PL1_A2" : DInt AT PosiciónEntrega_PL1(Ant), 1 s
   "PosiciónEntrega_PL2_A2" : DInt AT PosiciónEntrega_PL2(Ant), 1 s
   "PosiciónEspera_PL1_A2" : DInt AT PosiciónEspera_PL1(Ant), 1 s
   "PosiciónEspera_PL2_A2" : DInt AT PosiciónEspera_PL2(Ant), 1 s
   "PosiciónPlegado1_PL1_A2" : DInt AT PosiciónPlegado1_PL1(Ant), 1 s
   "PosiciónPlegado1_PL2_A2" : DInt AT PosiciónPlegado1_PL2(Ant), 1 s
   "PosiciónPlegado2_PL1_A2" : DInt AT PosiciónPlegado2_PL1(Ant), 1 s
   "PosiciónPlegado2_PL2_A2" : DInt AT PosiciónPlegado2_PL2(Ant), 1 s
   "PosiciónRecepción_PL1_A2" : DInt AT PosiciónRecepción_PL1(Ant), 1 s
   "PosiciónRecepción_PL2_A2" : DInt AT PosiciónRecepción_PL2(Ant), 1 s

graphic list "General - Plegadora": 0..1 'Plegador 1 G'; 1 'Plegador 2_1'

graphic list "General - Almacén": 0..1 'Almacen 1 G'; 1 'Almacen 2_1'

graphic list "General - Formador": 0..1 'F1_G'; 1 'F1R'

graphic list "General - Pinza": 0..1 'Pinza G'; 1 'Pinza 2_1'

graphic list "General - Cinta": 0..1 'Cinta G'; 1 'Cinta 2_1'

graphic list "General - Perfiladores": 0..1 'Perfiladores 1 G'; 1 'Perfiladores 2_1'

graphic list "General - Rolos": 0..1 'Rolos 1 G'; 1 'Rolos 2_3'

graphic list "General - Araña": 0..1 'Araña 1 G'; 1 'Araña 2_1'

graphic list "General - Descargador": 0..1 'Descargador G'; 1 'Descargador 2_1'

graphic list "GeneralBase": 0 'Base G'; 1 'BaseRoja'

screen "Principal" 1366x768, template "Template"
   GraphicIOField "Campo ES gráfico_10" at 43,115 size 1272x557; PictureList "GeneralBase"
      ProcessValue <- "Aux2"
   Button "Botón_13" at 1056,519 size 200x40; TextOff 'Limpiar Fichero'
      ObjectEnable <- "Aux3"
      Appearance <- "Aux3"
      on Press: function_ff1151d2(0, "FV_DatProducto_Alm1_"); function_ff1151d2(0, "FV_PosPinza_Alm1_"); function_ff1151d2(0, "FV_PosPlegadores_Alm1_"); function_ff1151d2(0, "FV_DatProducto_Alm2_"); function_ff1151d2(0, "FV_PosPinza_Alm2_"); function_ff1151d2(0, "FV_PosPlegadores_Alm2_"); function_ff1151d2(0, "FV_Defectos_Alm1_"); function_ff1151d2(0, "FV_Defectos_Alm2_")
   Button "Botón_11" at 1056,576 size 200x40; TextOff 'Detener archivado'
      on Click: function_efd5fb8c(); SetBit("Aux3")
      ObjectEnable <- "Aux3"
      Appearance <- "Aux3"
   Button "Botón_12" at 1056,633 size 200x40; TextOff 'Exportar archivos al Pendrive'
      Appearance <- "Aux3"
      on Press: function_e9be9208(0, "FV_DatProducto_Alm1_", 'D:\Roll Forming\Amacén 1', 0); function_e9be9208(0, "FV_PosPinza_Alm1_", 'D:\Roll Forming\Amacén 1', 0); function_e9be9208(0, "FV_PosPlegadores_Alm1_", 'D:\Roll Forming\Amacén 1', 0); function_e9be9208(0, "FV_DatProducto_Alm2_", 'D:\Roll Forming\Amacén 2', 0); function_e9be9208(0, "FV_PosPinza_Alm2_", 'D:\Roll Forming\Amacén 2', 0); function_e9be9208(0, "FV_PosPlegadores_Alm2_", 'D:\Roll Forming\Amacén 2', 0); function_e9be9208(0, "FV_Defectos_Alm1_", 'D:\Roll Forming\Amacén 1', 0); function_e9be9208(0, "FV_Defectos_Alm2_", 'D:\Roll Forming\Amacén 2', 0)
      ObjectEnable <- "Aux3"
   GraphicIOField "Campo ES gráfico_7" at 867,122 size 309x174; PictureList "General - Plegadora"
      ProcessValue <- "Aux2"
   GraphicIOField "Campo ES gráfico_2" at 98,389 size 219x150; PictureList "General - Almacén"
      ProcessValue <- "Aux2"
   GraphicIOField "Campo ES gráfico_8" at 798,281 size 77x78; PictureList "General - Formador"
      ProcessValue <- "Aux2"
   GraphicIOField "Campo ES gráfico_6" at 914,210 size 309x150; PictureList "General - Pinza"
      ProcessValue <- "Aux2"
   GraphicIOField "Campo ES gráfico_5" at 650,307 size 293x150; PictureList "General - Cinta"
      ProcessValue <- "Aux2"
   GraphicIOField "Campo ES gráfico_4" at 453,391 size 221x134; PictureList "General - Perfiladores"
      ProcessValue <- "Aux2"
   GraphicIOField "Campo ES gráfico_3" at 188,463 size 285x158; PictureList "General - Rolos"
      ProcessValue <- "Aux2"
   GraphicIOField "Campo ES gráfico_1" at 86,348 size 300x302; PictureList "General - Araña"
      ProcessValue <- "Aux2"
   GraphicIOField "Campo ES gráfico_9" at 1056,165 size 141x246; PictureList "General - Descargador"
      ProcessValue <- "Aux2"
   TextField "Campo de texto_1" at 36,62 size 465x92; Text 'Roll Forming'
   TextField "Campo de texto_28" at 35,249 size 65x20; Text 'Almacén 2'
   TextField "Campo de texto_29" at 35,209 size 65x20; Text 'Almacén 1'
   Button "Botón_31" at 0,697 size 137x70; TextOff 'Principal'
   IOField "Campo ES_2" at 313,203 size 96x32; FormatPattern 999999
      ProcessValue <- "Contador_def_Alm1"
   IOField "Campo ES_3" at 313,243 size 96x32; FormatPattern 999999
      ProcessValue <- "Contador_def_Alm2"
   TextField "Campo de texto_300" at 299,177 size 127x20; Text 'Contador de defectos'
   Button "Botón_10" at 1056,463 size 200x40; TextOff 'Iniciar archivado'
      on Release: function_bb0abc73(); function_fd9437ed(0, "FV_DatProducto_Alm1_"); function_fd9437ed(0, "FV_PosPinza_Alm1_"); function_fd9437ed(0, "FV_PosPlegadores_Alm1_"); function_fd9437ed(0, "FV_DatProducto_Alm2_"); function_fd9437ed(0, "FV_PosPinza_Alm2_"); function_fd9437ed(0, "FV_PosPlegadores_Alm2_"); function_fd9437ed(0, "FV_Defectos_Alm1_"); function_fd9437ed(0, "FV_Defectos_Alm2_"); ResetBit("Aux3")
      Appearance <- "Aux3"
      ObjectEnable <- "Aux3"
   Circle "Cercle_10" at 780,599 size 10x10
      Appearance <- "31S1 (E8.0)"
   Circle "Cercle_1" at 780,567 size 10x10
      Appearance <- "Descargador-PiezaPresente"
   TextField "Campo de texto_2" at 803,562 size 196x20; Text 'Pieza presente en el descargador'
   TextField "Campo de texto_3" at 803,594 size 34x20; Text '31S1'
   IOField "Champ E/S_57" at 123,246 size 118x24; FormatPattern ????????????????????
      ProcessValue <- "Almacén 2\PAlmacén.Nombre"
   IOField "Champ E/S_56" at 123,206 size 120x24; FormatPattern ????????????????????
      ProcessValue <- "Almacén 1\PAlmacén.Nombre"

Template "Template" 1366x768
   Button "Plantilla_Botón_2" at 689,697 size 552x70; TextOff 'Almacen 2'
   Button "Plantilla_Botón_1" at 137,697 size 552x70; TextOff 'Almacen 1'
   GraphicView "Visor de gráficos_3" at 78,7 size 94x30; Picture "eProC_B0"
   GraphicView "Visor de gráficos_4" at 20,7 size 53x30; Picture "eProC_A0"
   Button "Botón_1" at 276,725 size 137x40; TextOff 'Pos. de Pinza'
   Button "Botón_2" at 139,725 size 137x40; TextOff 'Factor "F"'
   Button "Botón_4" at 413,725 size 137x40; TextOff 'Factor "PL"'
   Button "Botón_5" at 550,725 size 137x40; TextOff 'Pos. de Pleg.'
   Button "Botón_3" at 0,697 size 137x70; TextOff 'Principal'
      on Click: ActivateScreen("Principal", 0)
   Button "Botón_6" at 828,725 size 137x40; TextOff 'Pos. de Pinza'
   Button "Botón_7" at 691,725 size 137x40; TextOff 'Factor "F"'
   Button "Botón_8" at 965,725 size 137x40; TextOff 'Factor "PL"'
   Button "Botón_9" at 1102,725 size 137x40; TextOff 'Pos. de Pleg.'
   Button "Plantilla_Botón_41" at 1241,697 size 125x70; TextOff 'Salir del runtime'
      on Press: StopRuntime(0)

VB script "FuncionVB_1"
   'Sugerencia:
   ' 1. Utilice la combinación de teclas <CTRL+ESPACIO> o <CTRL+I> para abrir una lista de todos los objetos y funciones
   ' 2. Escriba el código utilizando el objeto HMI Runtime.
   '  Ejemplo: HmiRuntime.Screens("Screen_1").
   ' 3. Utilice la combinación de teclas <CTRL+J> para crear una referencia de objeto..
   'Escriba el código a partir de esta posición:
   
   
   'Si hay pieza presente en el descargador
   If SmartTags("Descargador-PiezaPresente")=True Then
   	'y el sensor a la salida lee la unidad (descargador posiciòn atras)
   	If SmartTags("31S1 (E8.0)")=False Then 'And SmartTags("Aux1")=False , para guardar solo con el flanco ascendente de 31S1
   		'dependiendo de que almacen proviene (0=almacen 1; 1=almacen 2), conmuto la variable local que dispara el evento para guardar los datos en el fichero correspondiente
   		If SmartTags("Descargador-Almacen")=False Then
   			cd43ef6d-4af9-40c6-aa76-7baaf5848e36 Evento_ArchivarVariable_1
   			cd43ef6d-4af9-40c6-aa76-7baaf5848e36 Evento_ArchivarVariable_2
   			cd43ef6d-4af9-40c6-aa76-7baaf5848e36 Evento_ArchivarVariable_3
   		Else
   			cd43ef6d-4af9-40c6-aa76-7baaf5848e36 Evento_ArchivarVariable_4
   			cd43ef6d-4af9-40c6-aa76-7baaf5848e36 Evento_ArchivarVariable_5
   			cd43ef6d-4af9-40c6-aa76-7baaf5848e36 Evento_ArchivarVariable_6
   		End If
   		'SmartTags("Aux1")=True
   	End If
   Else
   'SmartTags("Aux1")=False
   End If
*)